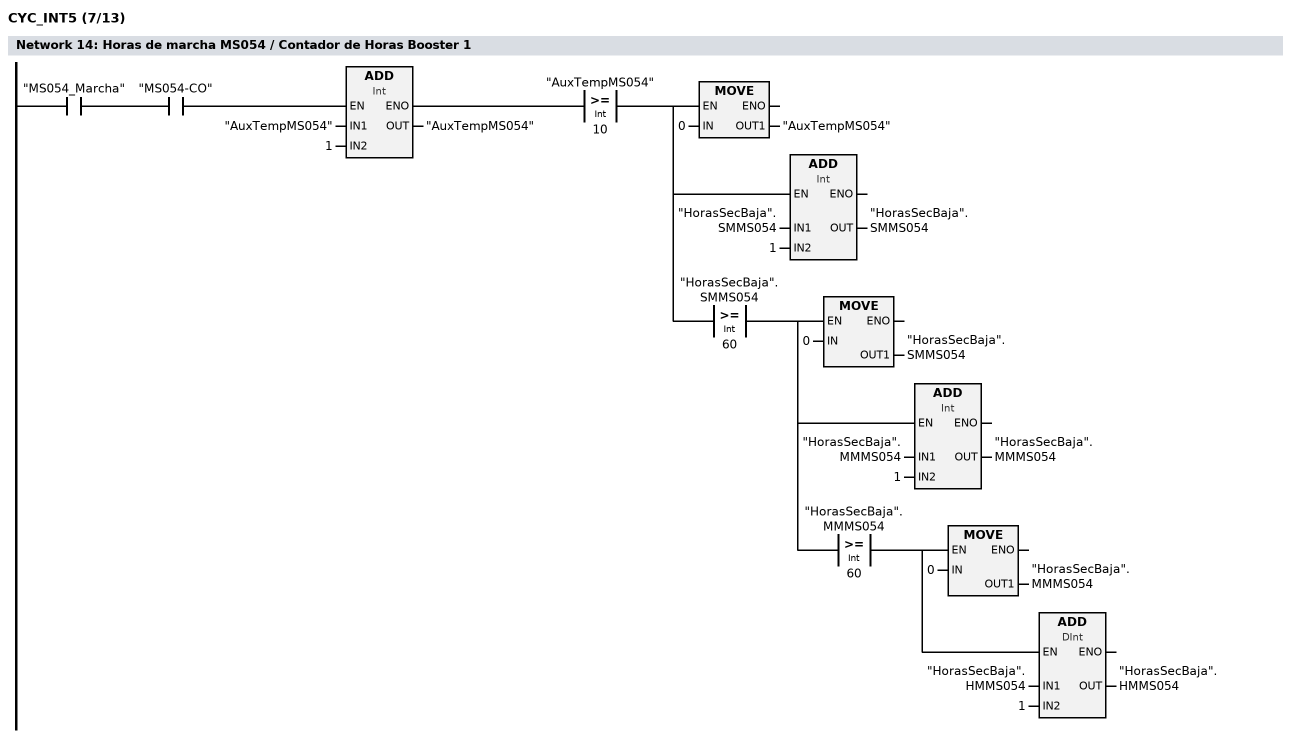
   RUNG wire#powerrail
      Contact( "MS054_Marcha" )
      Contact( "MS054-CO" )
      { S7_Templates := "SrcType := Int"; S7_GenerateENO := "TRUE" } Add(in1 := "AuxTempMS054", in2 := 1, out => "AuxTempMS054")
      { S7_Templates := "SrcType := Int" } GE_Contact(in1 := "AuxTempMS054", in2 := 10)
      wire#w1
      { S7_GenerateENO := "TRUE" } Move(in := 0, out1 => "AuxTempMS054")
   END_RUNG
   RUNG wire#w1
      { S7_Templates := "SrcType := Int"; S7_GenerateENO := "TRUE" } Add(in1 := "HorasSecBaja".SMMS054, in2 := 1, out => "HorasSecBaja".SMMS054)
   END_RUNG
   RUNG wire#w1
      { S7_Templates := "SrcType := Int" } GE_Contact(in1 := "HorasSecBaja".SMMS054, in2 := 60)
      wire#w2
      { S7_GenerateENO := "TRUE" } Move(in := 0, out1 => "HorasSecBaja".SMMS054)
   END_RUNG
   RUNG wire#w2
      { S7_Templates := "SrcType := Int"; S7_GenerateENO := "TRUE" } Add(in1 := "HorasSecBaja".MMMS054, in2 := 1, out => "HorasSecBaja".MMMS054)
   END_RUNG
   RUNG wire#w2
      { S7_Templates := "SrcType := Int" } GE_Contact(in1 := "HorasSecBaja".MMMS054, in2 := 60)
      wire#w3
      { S7_GenerateENO := "TRUE" } Move(in := 0, out1 => "HorasSecBaja".MMMS054)
   END_RUNG
   RUNG wire#w3
      { S7_Templates := "SrcType := DInt"; S7_GenerateENO := "TRUE" } Add(in1 := "HorasSecBaja".HMMS054, in2 := 1, out => "HorasSecBaja".HMMS054)
   END_RUNG
   // the same network as SCL:
   // ENO of a box is taken as its EN; it also drops when the box reports an error
   #_w1 := "MS054_Marcha" AND "MS054-CO";
   IF #_w1 THEN "AuxTempMS054" := "AuxTempMS054" + 1; END_IF;
   #_w2 := #_w1 AND ("AuxTempMS054" >= 10);
   IF #_w2 THEN
       "AuxTempMS054" := 0;
       "HorasSecBaja".SMMS054 := "HorasSecBaja".SMMS054 + 1;
   END_IF;
   #_w3 := #_w2 AND ("HorasSecBaja".SMMS054 >= 60);
   IF #_w3 THEN
       "HorasSecBaja".SMMS054 := 0;
       "HorasSecBaja".MMMS054 := "HorasSecBaja".MMMS054 + 1;
   END_IF;
   #_w4 := #_w3 AND ("HorasSecBaja".MMMS054 >= 60);
   IF #_w4 THEN
       "HorasSecBaja".MMMS054 := 0;
       "HorasSecBaja".HMMS054 := "HorasSecBaja".HMMS054 + 1;
   END_IF;
END_REGION

REGION Network 15: Horas de marcha MS055 / Contador de Horas Booster 1
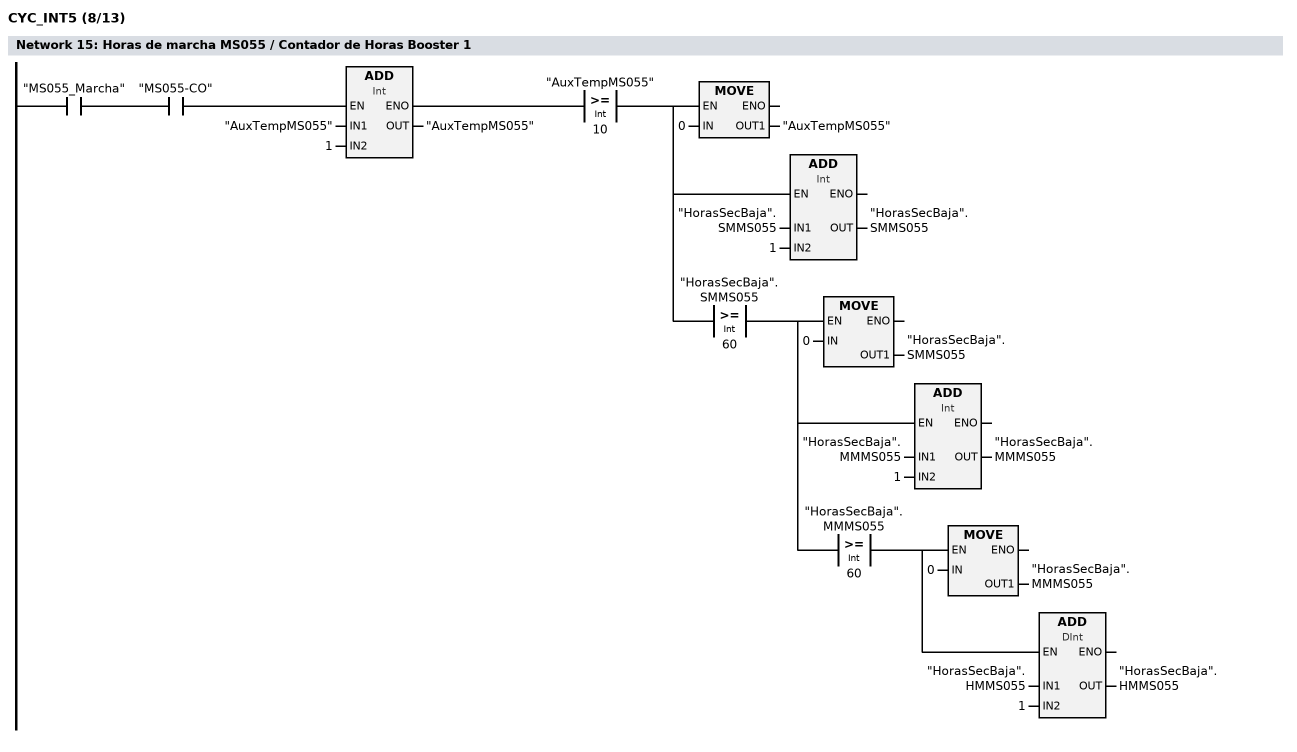
   RUNG wire#powerrail
      Contact( "MS055_Marcha" )
      Contact( "MS055-CO" )
      { S7_Templates := "SrcType := Int"; S7_GenerateENO := "TRUE" } Add(in1 := "AuxTempMS055", in2 := 1, out => "AuxTempMS055")
      { S7_Templates := "SrcType := Int" } GE_Contact(in1 := "AuxTempMS055", in2 := 10)
      wire#w1
      { S7_GenerateENO := "TRUE" } Move(in := 0, out1 => "AuxTempMS055")
   END_RUNG
   RUNG wire#w1
      { S7_Templates := "SrcType := Int"; S7_GenerateENO := "TRUE" } Add(in1 := "HorasSecBaja".SMMS055, in2 := 1, out => "HorasSecBaja".SMMS055)
   END_RUNG
   RUNG wire#w1
      { S7_Templates := "SrcType := Int" } GE_Contact(in1 := "HorasSecBaja".SMMS055, in2 := 60)
      wire#w2
      { S7_GenerateENO := "TRUE" } Move(in := 0, out1 => "HorasSecBaja".SMMS055)
   END_RUNG
   RUNG wire#w2
      { S7_Templates := "SrcType := Int"; S7_GenerateENO := "TRUE" } Add(in1 := "HorasSecBaja".MMMS055, in2 := 1, out => "HorasSecBaja".MMMS055)
   END_RUNG
   RUNG wire#w2
      { S7_Templates := "SrcType := Int" } GE_Contact(in1 := "HorasSecBaja".MMMS055, in2 := 60)
      wire#w3
      { S7_GenerateENO := "TRUE" } Move(in := 0, out1 => "HorasSecBaja".MMMS055)
   END_RUNG
   RUNG wire#w3
      { S7_Templates := "SrcType := DInt"; S7_GenerateENO := "TRUE" } Add(in1 := "HorasSecBaja".HMMS055, in2 := 1, out => "HorasSecBaja".HMMS055)
   END_RUNG
   // the same network as SCL:
   // ENO of a box is taken as its EN; it also drops when the box reports an error
   #_w1 := "MS055_Marcha" AND "MS055-CO";
   IF #_w1 THEN "AuxTempMS055" := "AuxTempMS055" + 1; END_IF;
   #_w2 := #_w1 AND ("AuxTempMS055" >= 10);
   IF #_w2 THEN
       "AuxTempMS055" := 0;
       "HorasSecBaja".SMMS055 := "HorasSecBaja".SMMS055 + 1;
   END_IF;
   #_w3 := #_w2 AND ("HorasSecBaja".SMMS055 >= 60);
   IF #_w3 THEN
       "HorasSecBaja".SMMS055 := 0;
       "HorasSecBaja".MMMS055 := "HorasSecBaja".MMMS055 + 1;
   END_IF;
   #_w4 := #_w3 AND ("HorasSecBaja".MMMS055 >= 60);
   IF #_w4 THEN
       "HorasSecBaja".MMMS055 := 0;
       "HorasSecBaja".HMMS055 := "HorasSecBaja".HMMS055 + 1;
   END_IF;
END_REGION

REGION Network 16: Horas de marcha MC060 / Contador de Horas Booster 1
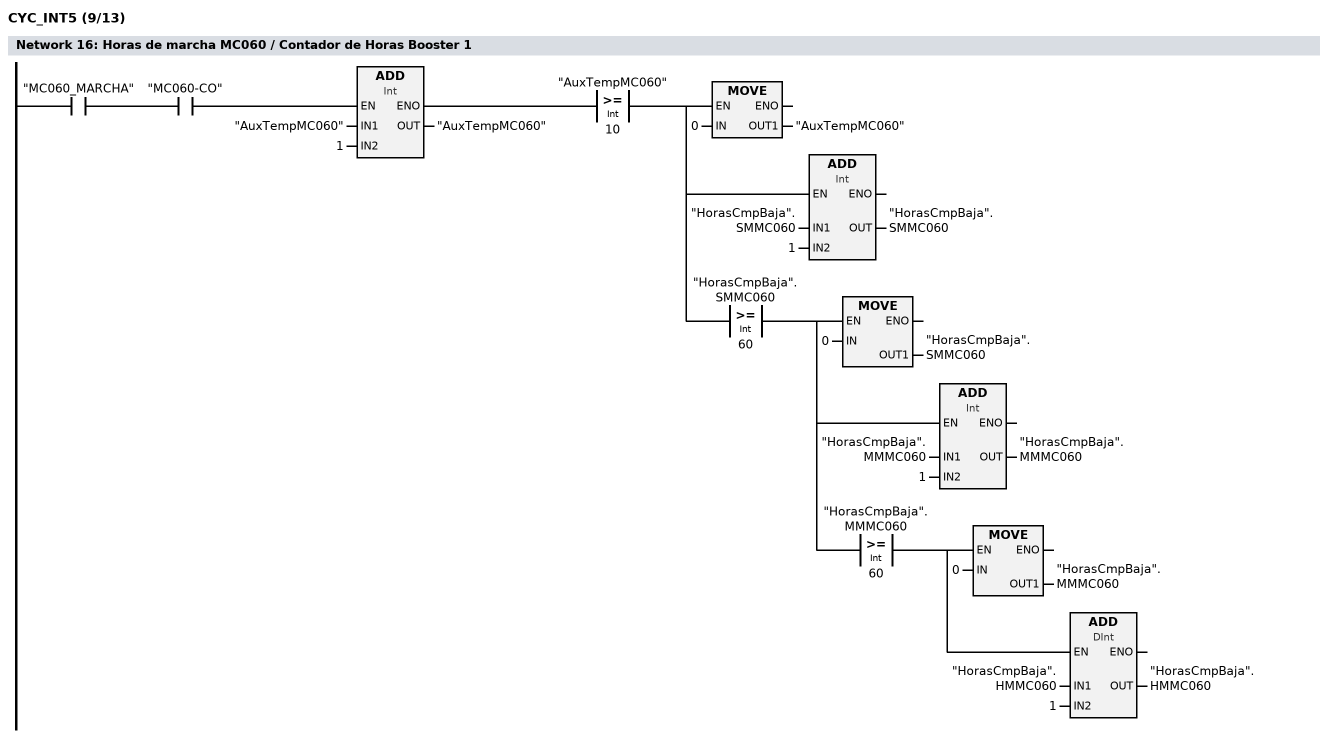
   RUNG wire#powerrail
      Contact( "MC060_MARCHA" )
      Contact( "MC060-CO" )
      { S7_Templates := "SrcType := Int"; S7_GenerateENO := "TRUE" } Add(in1 := "AuxTempMC060", in2 := 1, out => "AuxTempMC060")
      { S7_Templates := "SrcType := Int" } GE_Contact(in1 := "AuxTempMC060", in2 := 10)
      wire#w1
      { S7_GenerateENO := "TRUE" } Move(in := 0, out1 => "AuxTempMC060")
   END_RUNG
   RUNG wire#w1
      { S7_Templates := "SrcType := Int"; S7_GenerateENO := "TRUE" } Add(in1 := "HorasCmpBaja".SMMC060, in2 := 1, out => "HorasCmpBaja".SMMC060)
   END_RUNG
   RUNG wire#w1
      { S7_Templates := "SrcType := Int" } GE_Contact(in1 := "HorasCmpBaja".SMMC060, in2 := 60)
      wire#w2
      { S7_GenerateENO := "TRUE" } Move(in := 0, out1 => "HorasCmpBaja".SMMC060)
   END_RUNG
   RUNG wire#w2
      { S7_Templates := "SrcType := Int"; S7_GenerateENO := "TRUE" } Add(in1 := "HorasCmpBaja".MMMC060, in2 := 1, out => "HorasCmpBaja".MMMC060)
   END_RUNG
   RUNG wire#w2
      { S7_Templates := "SrcType := Int" } GE_Contact(in1 := "HorasCmpBaja".MMMC060, in2 := 60)
      wire#w3
      { S7_GenerateENO := "TRUE" } Move(in := 0, out1 => "HorasCmpBaja".MMMC060)
   END_RUNG
   RUNG wire#w3
      { S7_Templates := "SrcType := DInt"; S7_GenerateENO := "TRUE" } Add(in1 := "HorasCmpBaja".HMMC060, in2 := 1, out => "HorasCmpBaja".HMMC060)
   END_RUNG
   // the same network as SCL:
   // ENO of a box is taken as its EN; it also drops when the box reports an error
   #_w1 := "MC060_MARCHA" AND "MC060-CO";
   IF #_w1 THEN "AuxTempMC060" := "AuxTempMC060" + 1; END_IF;
   #_w2 := #_w1 AND ("AuxTempMC060" >= 10);
   IF #_w2 THEN
       "AuxTempMC060" := 0;
       "HorasCmpBaja".SMMC060 := "HorasCmpBaja".SMMC060 + 1;
   END_IF;
   #_w3 := #_w2 AND ("HorasCmpBaja".SMMC060 >= 60);
   IF #_w3 THEN
       "HorasCmpBaja".SMMC060 := 0;
       "HorasCmpBaja".MMMC060 := "HorasCmpBaja".MMMC060 + 1;
   END_IF;
   #_w4 := #_w3 AND ("HorasCmpBaja".MMMC060 >= 60);
   IF #_w4 THEN
       "HorasCmpBaja".MMMC060 := 0;
       "HorasCmpBaja".HMMC060 := "HorasCmpBaja".HMMC060 + 1;
   END_IF;
END_REGION

REGION Network 17: Horas de marcha MC061 / Contador de Horas Booster 1
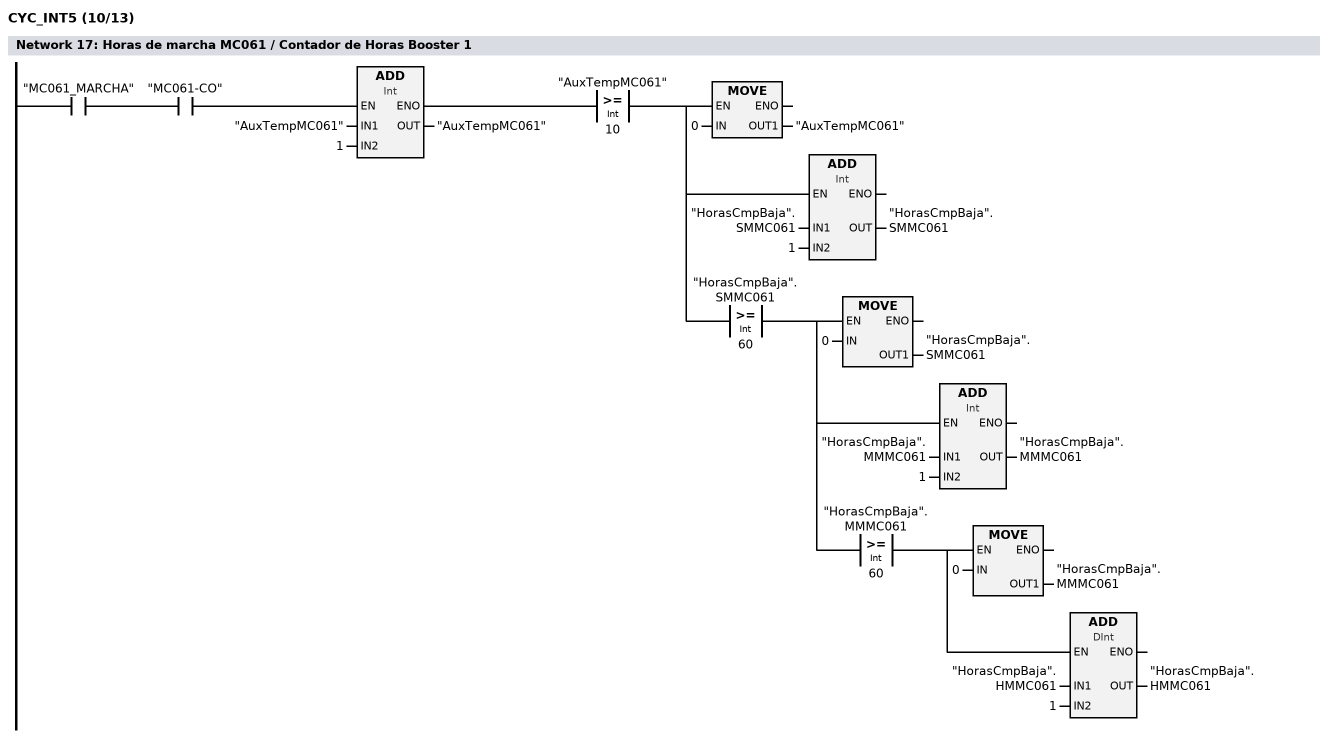
   RUNG wire#powerrail
      Contact( "MC061_MARCHA" )
      Contact( "MC061-CO" )
      { S7_Templates := "SrcType := Int"; S7_GenerateENO := "TRUE" } Add(in1 := "AuxTempMC061", in2 := 1, out => "AuxTempMC061")
      { S7_Templates := "SrcType := Int" } GE_Contact(in1 := "AuxTempMC061", in2 := 10)
      wire#w1
      { S7_GenerateENO := "TRUE" } Move(in := 0, out1 => "AuxTempMC061")
   END_RUNG
   RUNG wire#w1
      { S7_Templates := "SrcType := Int"; S7_GenerateENO := "TRUE" } Add(in1 := "HorasCmpBaja".SMMC061, in2 := 1, out => "HorasCmpBaja".SMMC061)
   END_RUNG
   RUNG wire#w1
      { S7_Templates := "SrcType := Int" } GE_Contact(in1 := "HorasCmpBaja".SMMC061, in2 := 60)
      wire#w2
      { S7_GenerateENO := "TRUE" } Move(in := 0, out1 => "HorasCmpBaja".SMMC061)
   END_RUNG
   RUNG wire#w2
      { S7_Templates := "SrcType := Int"; S7_GenerateENO := "TRUE" } Add(in1 := "HorasCmpBaja".MMMC061, in2 := 1, out => "HorasCmpBaja".MMMC061)
   END_RUNG
   RUNG wire#w2
      { S7_Templates := "SrcType := Int" } GE_Contact(in1 := "HorasCmpBaja".MMMC061, in2 := 60)
      wire#w3
      { S7_GenerateENO := "TRUE" } Move(in := 0, out1 => "HorasCmpBaja".MMMC061)
   END_RUNG
   RUNG wire#w3
      { S7_Templates := "SrcType := DInt"; S7_GenerateENO := "TRUE" } Add(in1 := "HorasCmpBaja".HMMC061, in2 := 1, out => "HorasCmpBaja".HMMC061)
   END_RUNG
   // the same network as SCL:
   // ENO of a box is taken as its EN; it also drops when the box reports an error
   #_w1 := "MC061_MARCHA" AND "MC061-CO";
   IF #_w1 THEN "AuxTempMC061" := "AuxTempMC061" + 1; END_IF;
   #_w2 := #_w1 AND ("AuxTempMC061" >= 10);
   IF #_w2 THEN
       "AuxTempMC061" := 0;
       "HorasCmpBaja".SMMC061 := "HorasCmpBaja".SMMC061 + 1;
   END_IF;
   #_w3 := #_w2 AND ("HorasCmpBaja".SMMC061 >= 60);
   IF #_w3 THEN
       "HorasCmpBaja".SMMC061 := 0;
       "HorasCmpBaja".MMMC061 := "HorasCmpBaja".MMMC061 + 1;
   END_IF;
   #_w4 := #_w3 AND ("HorasCmpBaja".MMMC061 >= 60);
   IF #_w4 THEN
       "HorasCmpBaja".MMMC061 := 0;
       "HorasCmpBaja".HMMC061 := "HorasCmpBaja".HMMC061 + 1;
   END_IF;
END_REGION

REGION Network 18: Horas de marcha MC062 / Contador de Horas Booster 1
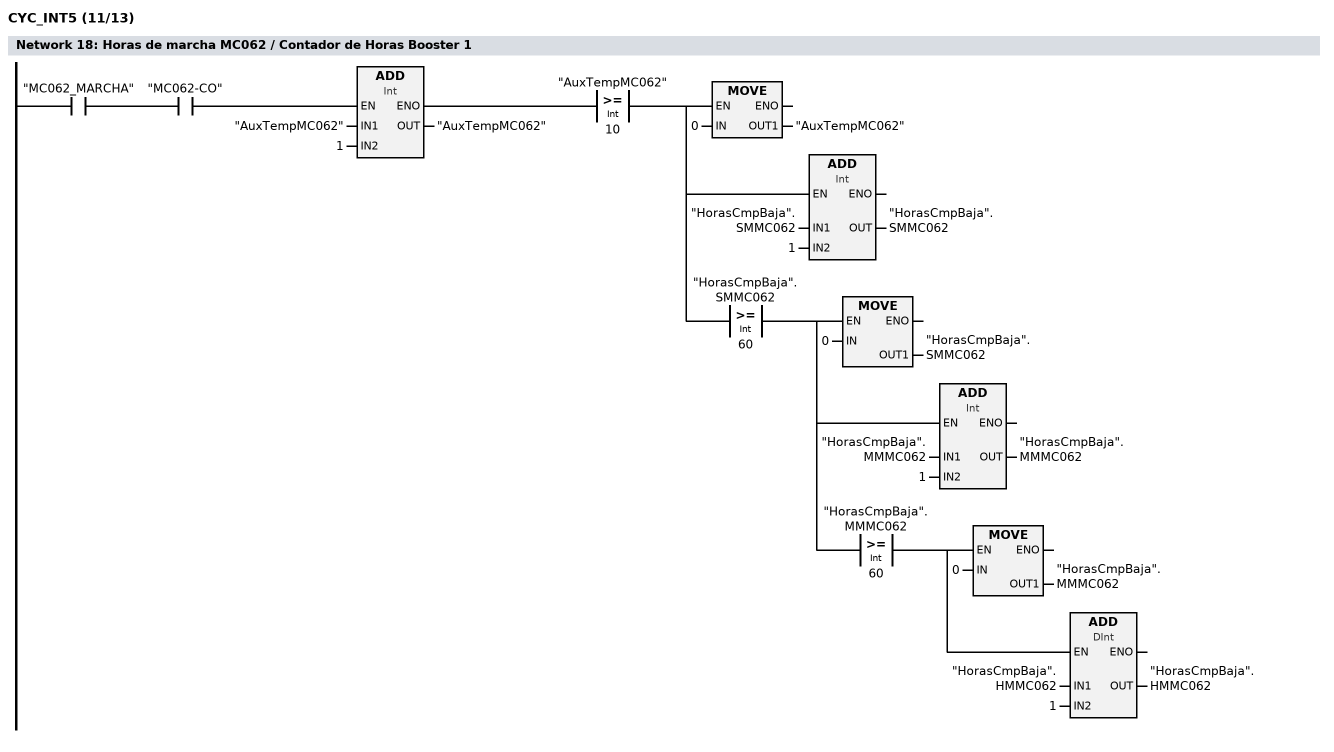
   RUNG wire#powerrail
      Contact( "MC062_MARCHA" )
      Contact( "MC062-CO" )
      { S7_Templates := "SrcType := Int"; S7_GenerateENO := "TRUE" } Add(in1 := "AuxTempMC062", in2 := 1, out => "AuxTempMC062")
      { S7_Templates := "SrcType := Int" } GE_Contact(in1 := "AuxTempMC062", in2 := 10)
      wire#w1
      { S7_GenerateENO := "TRUE" } Move(in := 0, out1 => "AuxTempMC062")
   END_RUNG
   RUNG wire#w1
      { S7_Templates := "SrcType := Int"; S7_GenerateENO := "TRUE" } Add(in1 := "HorasCmpBaja".SMMC062, in2 := 1, out => "HorasCmpBaja".SMMC062)
   END_RUNG
   RUNG wire#w1
      { S7_Templates := "SrcType := Int" } GE_Contact(in1 := "HorasCmpBaja".SMMC062, in2 := 60)
      wire#w2
      { S7_GenerateENO := "TRUE" } Move(in := 0, out1 => "HorasCmpBaja".SMMC062)
   END_RUNG
   RUNG wire#w2
      { S7_Templates := "SrcType := Int"; S7_GenerateENO := "TRUE" } Add(in1 := "HorasCmpBaja".MMMC062, in2 := 1, out => "HorasCmpBaja".MMMC062)
   END_RUNG
   RUNG wire#w2
      { S7_Templates := "SrcType := Int" } GE_Contact(in1 := "HorasCmpBaja".MMMC062, in2 := 60)
      wire#w3
      { S7_GenerateENO := "TRUE" } Move(in := 0, out1 => "HorasCmpBaja".MMMC062)
   END_RUNG
   RUNG wire#w3
      { S7_Templates := "SrcType := DInt"; S7_GenerateENO := "TRUE" } Add(in1 := "HorasCmpBaja".HMMC062, in2 := 1, out => "HorasCmpBaja".HMMC062)
   END_RUNG
   // the same network as SCL:
   // ENO of a box is taken as its EN; it also drops when the box reports an error
   #_w1 := "MC062_MARCHA" AND "MC062-CO";
   IF #_w1 THEN "AuxTempMC062" := "AuxTempMC062" + 1; END_IF;
   #_w2 := #_w1 AND ("AuxTempMC062" >= 10);
   IF #_w2 THEN
       "AuxTempMC062" := 0;
       "HorasCmpBaja".SMMC062 := "HorasCmpBaja".SMMC062 + 1;
   END_IF;
   #_w3 := #_w2 AND ("HorasCmpBaja".SMMC062 >= 60);
   IF #_w3 THEN
       "HorasCmpBaja".SMMC062 := 0;
       "HorasCmpBaja".MMMC062 := "HorasCmpBaja".MMMC062 + 1;
   END_IF;
   #_w4 := #_w3 AND ("HorasCmpBaja".MMMC062 >= 60);
   IF #_w4 THEN
       "HorasCmpBaja".MMMC062 := 0;
       "HorasCmpBaja".HMMC062 := "HorasCmpBaja".HMMC062 + 1;
   END_IF;
END_REGION

REGION Network 19: Horas de marcha MC063 / Contador de Horas Booster 1
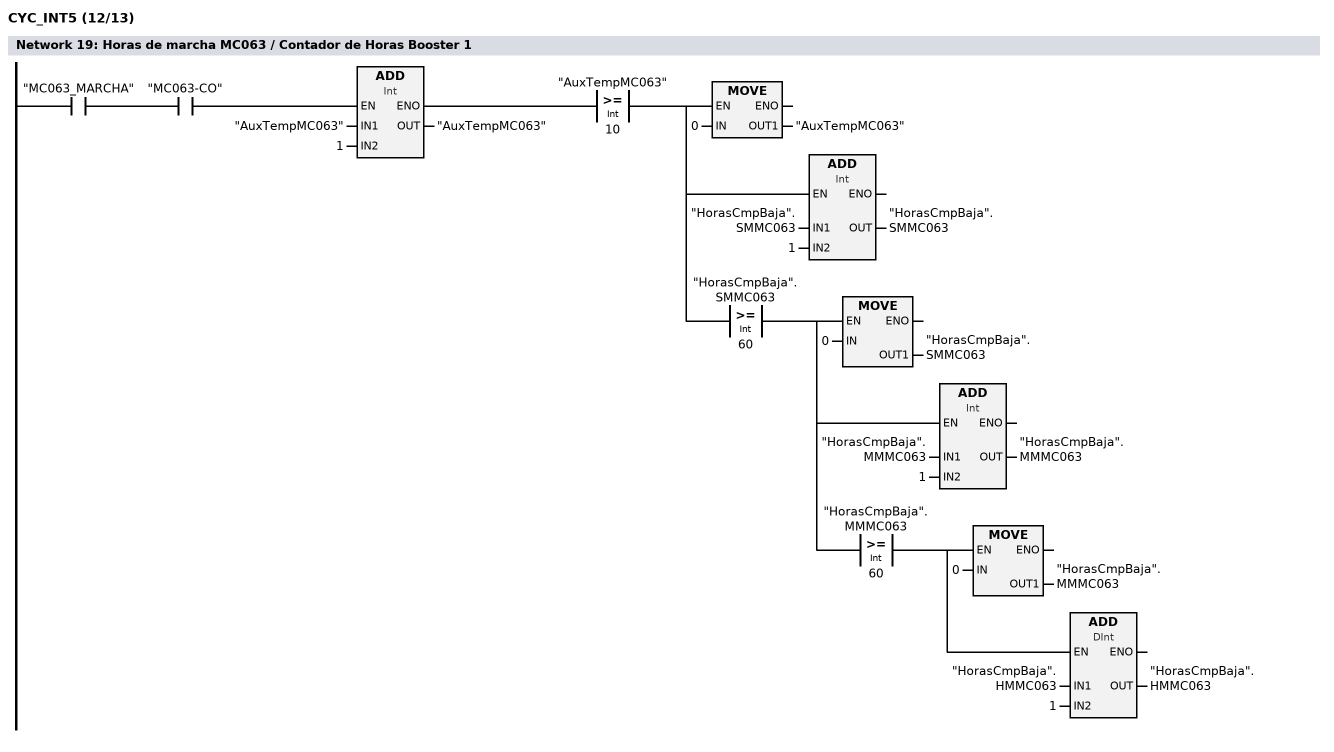
   RUNG wire#powerrail
      Contact( "MC063_MARCHA" )
      Contact( "MC063-CO" )
      { S7_Templates := "SrcType := Int"; S7_GenerateENO := "TRUE" } Add(in1 := "AuxTempMC063", in2 := 1, out => "AuxTempMC063")
      { S7_Templates := "SrcType := Int" } GE_Contact(in1 := "AuxTempMC063", in2 := 10)
      wire#w1
      { S7_GenerateENO := "TRUE" } Move(in := 0, out1 => "AuxTempMC063")
   END_RUNG
   RUNG wire#w1
      { S7_Templates := "SrcType := Int"; S7_GenerateENO := "TRUE" } Add(in1 := "HorasCmpBaja".SMMC063, in2 := 1, out => "HorasCmpBaja".SMMC063)
   END_RUNG
   RUNG wire#w1
      { S7_Templates := "SrcType := Int" } GE_Contact(in1 := "HorasCmpBaja".SMMC063, in2 := 60)
      wire#w2
      { S7_GenerateENO := "TRUE" } Move(in := 0, out1 => "HorasCmpBaja".SMMC063)
   END_RUNG
   RUNG wire#w2
      { S7_Templates := "SrcType := Int"; S7_GenerateENO := "TRUE" } Add(in1 := "HorasCmpBaja".MMMC063, in2 := 1, out => "HorasCmpBaja".MMMC063)
   END_RUNG
   RUNG wire#w2
      { S7_Templates := "SrcType := Int" } GE_Contact(in1 := "HorasCmpBaja".MMMC063, in2 := 60)
      wire#w3
      { S7_GenerateENO := "TRUE" } Move(in := 0, out1 => "HorasCmpBaja".MMMC063)
   END_RUNG
   RUNG wire#w3
      { S7_Templates := "SrcType := DInt"; S7_GenerateENO := "TRUE" } Add(in1 := "HorasCmpBaja".HMMC063, in2 := 1, out => "HorasCmpBaja".HMMC063)
   END_RUNG
   // the same network as SCL:
   // ENO of a box is taken as its EN; it also drops when the box reports an error
   #_w1 := "MC063_MARCHA" AND "MC063-CO";
   IF #_w1 THEN "AuxTempMC063" := "AuxTempMC063" + 1; END_IF;
   #_w2 := #_w1 AND ("AuxTempMC063" >= 10);
   IF #_w2 THEN
       "AuxTempMC063" := 0;
       "HorasCmpBaja".SMMC063 := "HorasCmpBaja".SMMC063 + 1;
   END_IF;
   #_w3 := #_w2 AND ("HorasCmpBaja".SMMC063 >= 60);
   IF #_w3 THEN
       "HorasCmpBaja".SMMC063 := 0;
       "HorasCmpBaja".MMMC063 := "HorasCmpBaja".MMMC063 + 1;
   END_IF;
   #_w4 := #_w3 AND ("HorasCmpBaja".MMMC063 >= 60);
   IF #_w4 THEN
       "HorasCmpBaja".MMMC063 := 0;
       "HorasCmpBaja".HMMC063 := "HorasCmpBaja".HMMC063 + 1;
   END_IF;
END_REGION

REGION Network 20: Horas de marcha MC064 / Contador de Horas Booster 1
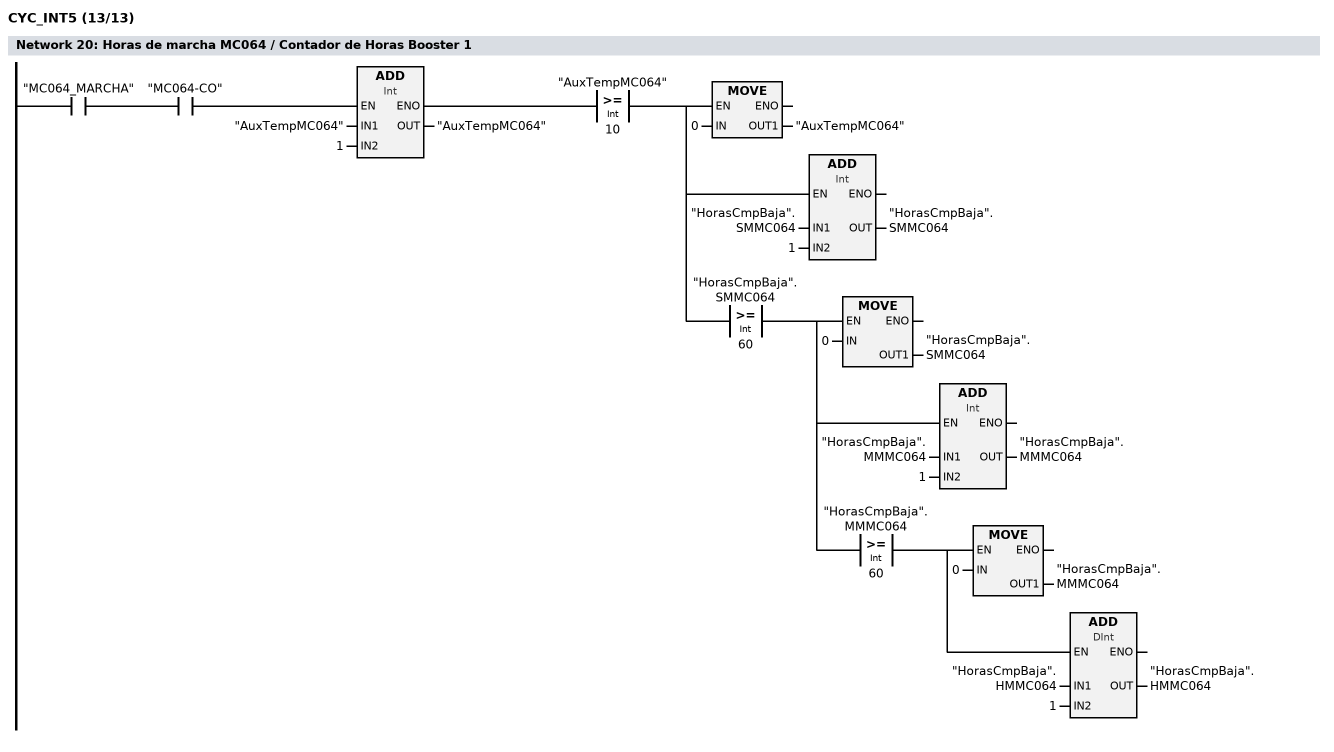
   RUNG wire#powerrail
      Contact( "MC064_MARCHA" )
      Contact( "MC064-CO" )
      { S7_Templates := "SrcType := Int"; S7_GenerateENO := "TRUE" } Add(in1 := "AuxTempMC064", in2 := 1, out => "AuxTempMC064")
      { S7_Templates := "SrcType := Int" } GE_Contact(in1 := "AuxTempMC064", in2 := 10)
      wire#w1
      { S7_GenerateENO := "TRUE" } Move(in := 0, out1 => "AuxTempMC064")
   END_RUNG
   RUNG wire#w1
      { S7_Templates := "SrcType := Int"; S7_GenerateENO := "TRUE" } Add(in1 := "HorasCmpBaja".SMMC064, in2 := 1, out => "HorasCmpBaja".SMMC064)
   END_RUNG
   RUNG wire#w1
      { S7_Templates := "SrcType := Int" } GE_Contact(in1 := "HorasCmpBaja".SMMC064, in2 := 60)
      wire#w2
      { S7_GenerateENO := "TRUE" } Move(in := 0, out1 => "HorasCmpBaja".SMMC064)
   END_RUNG
   RUNG wire#w2
      { S7_Templates := "SrcType := Int"; S7_GenerateENO := "TRUE" } Add(in1 := "HorasCmpBaja".MMMC064, in2 := 1, out => "HorasCmpBaja".MMMC064)
   END_RUNG
   RUNG wire#w2
      { S7_Templates := "SrcType := Int" } GE_Contact(in1 := "HorasCmpBaja".MMMC064, in2 := 60)
      wire#w3
      { S7_GenerateENO := "TRUE" } Move(in := 0, out1 => "HorasCmpBaja".MMMC064)
   END_RUNG
   RUNG wire#w3
      { S7_Templates := "SrcType := DInt"; S7_GenerateENO := "TRUE" } Add(in1 := "HorasCmpBaja".HMMC064, in2 := 1, out => "HorasCmpBaja".HMMC064)
   END_RUNG
   // the same network as SCL:
   // ENO of a box is taken as its EN; it also drops when the box reports an error
   #_w1 := "MC064_MARCHA" AND "MC064-CO";
   IF #_w1 THEN "AuxTempMC064" := "AuxTempMC064" + 1; END_IF;
   #_w2 := #_w1 AND ("AuxTempMC064" >= 10);
   IF #_w2 THEN
       "AuxTempMC064" := 0;
       "HorasCmpBaja".SMMC064 := "HorasCmpBaja".SMMC064 + 1;
   END_IF;
   #_w3 := #_w2 AND ("HorasCmpBaja".SMMC064 >= 60);
   IF #_w3 THEN
       "HorasCmpBaja".SMMC064 := 0;
       "HorasCmpBaja".MMMC064 := "HorasCmpBaja".MMMC064 + 1;
   END_IF;
   #_w4 := #_w3 AND ("HorasCmpBaja".MMMC064 >= 60);
   IF #_w4 THEN
       "HorasCmpBaja".MMMC064 := 0;
       "HorasCmpBaja".HMMC064 := "HorasCmpBaja".HMMC064 + 1;
   END_IF;
END_REGION
END_ORGANIZATION_BLOCK

// folder: OBs de Fallas

ORGANIZATION_BLOCK "OB40"   // OB40, STL
{ S7_Optimized_Access := 'FALSE' }
VERSION : 0.0
BEGIN
END_ORGANIZATION_BLOCK

ORGANIZATION_BLOCK "Cycle Time Fault"   // OB80, STL
{ S7_Optimized_Access := 'FALSE' }
VERSION : 0.0
BEGIN
END_ORGANIZATION_BLOCK

ORGANIZATION_BLOCK "I/O Point Fault 1"   // OB82, LAD
{ S7_Optimized_Access := 'FALSE' }
VERSION : 0.1
BEGIN
END_ORGANIZATION_BLOCK

ORGANIZATION_BLOCK "OB83"   // OB83, STL
{ S7_Optimized_Access := 'FALSE' }
VERSION : 0.1
BEGIN
END_ORGANIZATION_BLOCK

ORGANIZATION_BLOCK "OB Not Loaded Fault"   // OB85, LAD
{ S7_Optimized_Access := 'FALSE' }
VERSION : 0.1
BEGIN
END_ORGANIZATION_BLOCK

ORGANIZATION_BLOCK "Fallo del bastidor"   // OB86, STL
{ S7_Optimized_Access := 'FALSE' }
VERSION : 0.1
BEGIN
END_ORGANIZATION_BLOCK

ORGANIZATION_BLOCK "Communication Fault"   // OB87, LAD
{ S7_Optimized_Access := 'FALSE' }
VERSION : 0.1
BEGIN
END_ORGANIZATION_BLOCK

ORGANIZATION_BLOCK "Complete Restart"   // OB100, LAD
{ S7_Optimized_Access := 'FALSE' }
VERSION : 0.1
BEGIN
END_ORGANIZATION_BLOCK

ORGANIZATION_BLOCK "Programming Error"   // OB121, LAD
{ S7_Optimized_Access := 'FALSE' }
VERSION : 0.1
BEGIN
END_ORGANIZATION_BLOCK

ORGANIZATION_BLOCK "Module Access Error"   // OB122, LAD
{ S7_Optimized_Access := 'FALSE' }
VERSION : 0.1
BEGIN
END_ORGANIZATION_BLOCK

// folder: Panel

FUNCTION_BLOCK "CHControlMotorPanelMTA"   // FB55, LAD
{ S7_Optimized_Access := 'FALSE' }
VERSION : 0.1
   VAR_TEMP   // added for the SCL form of the ladder/FBD networks
      _w1 : Bool;
   END_VAR
BEGIN

REGION Network 1
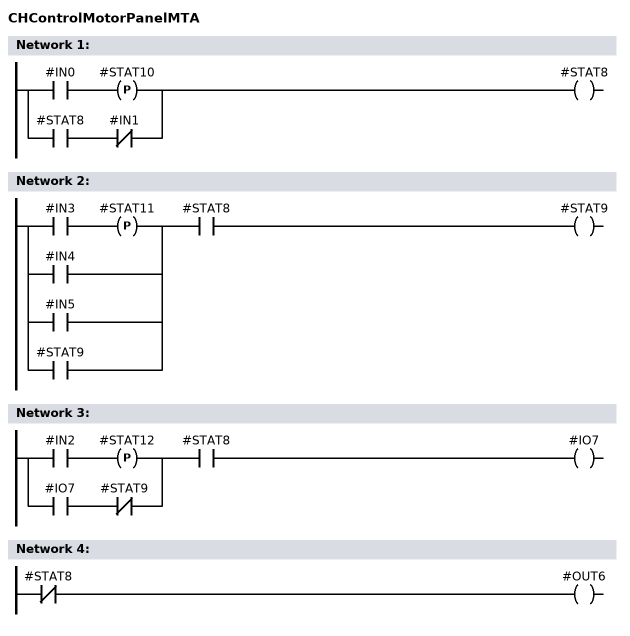
   RUNG wire#powerrail
      Contact( #IN0 )
      P_Trig( #STAT10 )
      wire#w1
      Coil( #STAT8 )
   END_RUNG
   RUNG wire#powerrail
      Contact( #STAT8 )
      I_Contact( #IN1 )
   END_RUNG wire#w1
   // the same network as SCL:
   #_w1 := #IN0 AND NOT #STAT10;   // rising edge
   #STAT10 := #IN0;
   #STAT8 := #_w1 OR (#STAT8 AND NOT #IN1);
END_REGION

REGION Network 2
   RUNG wire#powerrail
      Contact( #IN3 )
      P_Trig( #STAT11 )
      wire#w1
      Contact( #STAT8 )
      Coil( #STAT9 )
   END_RUNG
   RUNG wire#powerrail
      Contact( #IN4 )
   END_RUNG wire#w1
   RUNG wire#powerrail
      Contact( #IN5 )
   END_RUNG wire#w1
   RUNG wire#powerrail
      Contact( #STAT9 )
   END_RUNG wire#w1
   // the same network as SCL:
   #_w1 := #IN3 AND NOT #STAT11;   // rising edge
   #STAT11 := #IN3;
   #STAT9 := (#_w1 OR #IN4 OR #IN5 OR #STAT9) AND #STAT8;
END_REGION

REGION Network 3
   RUNG wire#powerrail
      Contact( #IN2 )
      P_Trig( #STAT12 )
      wire#w1
      Contact( #STAT8 )
      Coil( #IO7 )
   END_RUNG
   RUNG wire#powerrail
      Contact( #IO7 )
      I_Contact( #STAT9 )
   END_RUNG wire#w1
   // the same network as SCL:
   #_w1 := #IN2 AND NOT #STAT12;   // rising edge
   #STAT12 := #IN2;
   #IO7 := (#_w1 OR (#IO7 AND NOT #STAT9)) AND #STAT8;
END_REGION

REGION Network 4
   RUNG wire#powerrail
      I_Contact( #STAT8 )
      Coil( #OUT6 )
   END_RUNG
   // the same network as SCL:
   #OUT6 := NOT #STAT8;
END_REGION
END_FUNCTION_BLOCK

FUNCTION "AnimaciónMTA" : Void   // FC2, LAD
{ S7_Optimized_Access := 'FALSE' }
VERSION : 0.1
   VAR_TEMP   // added for the SCL form of the ladder/FBD networks
      _w1 : Bool;
      _w2 : Bool;
   END_VAR
BEGIN

REGION Network 1: Indicador Chillers
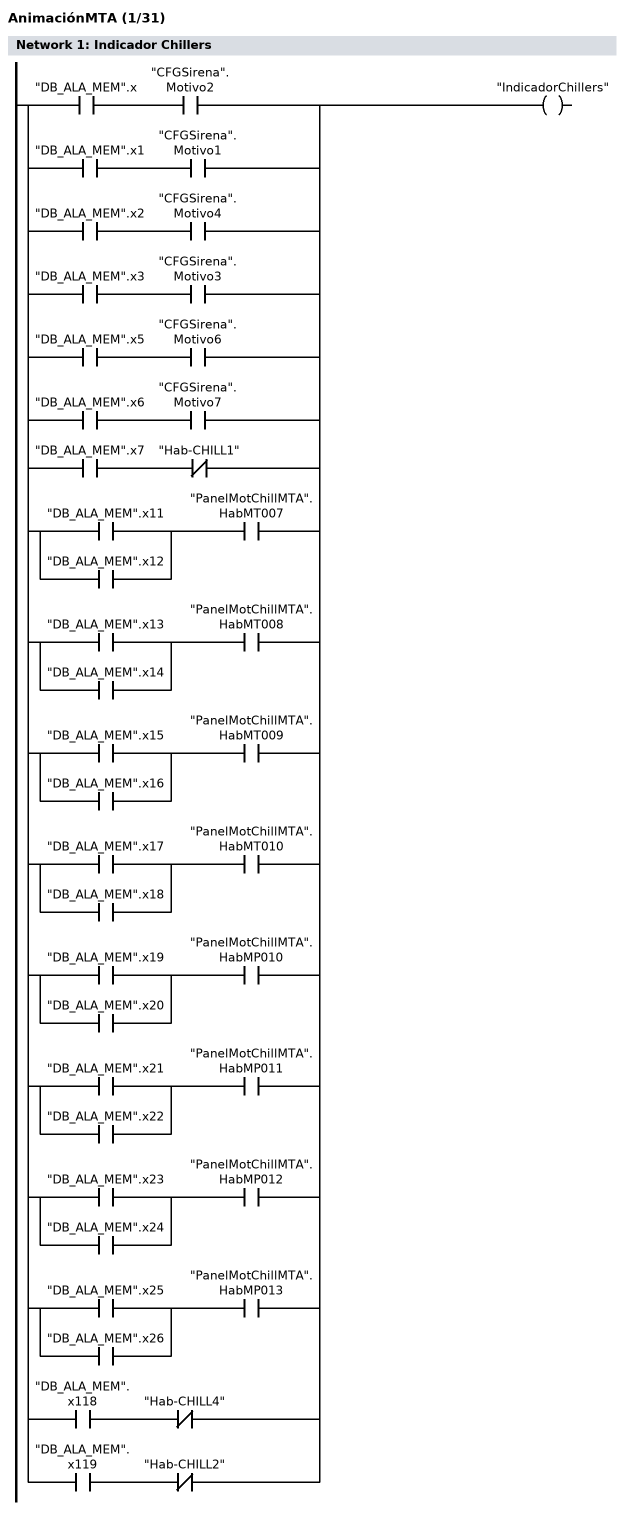
   RUNG wire#powerrail
      Contact( "DB_ALA_MEM".x )
      Contact( "CFGSirena".Motivo2 )
      wire#w1
      Coil( "IndicadorChillers" )
   END_RUNG
   RUNG wire#powerrail
      Contact( "DB_ALA_MEM".x1 )
      Contact( "CFGSirena".Motivo1 )
   END_RUNG wire#w1
   RUNG wire#powerrail
      Contact( "DB_ALA_MEM".x2 )
      Contact( "CFGSirena".Motivo4 )
   END_RUNG wire#w1
   RUNG wire#powerrail
      Contact( "DB_ALA_MEM".x3 )
      Contact( "CFGSirena".Motivo3 )
   END_RUNG wire#w1
   RUNG wire#powerrail
      Contact( "DB_ALA_MEM".x5 )
      Contact( "CFGSirena".Motivo6 )
   END_RUNG wire#w1
   RUNG wire#powerrail
      Contact( "DB_ALA_MEM".x6 )
      Contact( "CFGSirena".Motivo7 )
   END_RUNG wire#w1
   RUNG wire#powerrail
      Contact( "DB_ALA_MEM".x7 )
      I_Contact( "Hab-CHILL1" )
   END_RUNG wire#w1
   RUNG wire#powerrail
      Contact( "DB_ALA_MEM".x11 )
      wire#w2
      Contact( "PanelMotChillMTA".HabMT007 )
   END_RUNG wire#w1
   RUNG wire#powerrail
      Contact( "DB_ALA_MEM".x12 )
   END_RUNG wire#w2
   RUNG wire#powerrail
      Contact( "DB_ALA_MEM".x13 )
      wire#w3
      Contact( "PanelMotChillMTA".HabMT008 )
   END_RUNG wire#w1
   RUNG wire#powerrail
      Contact( "DB_ALA_MEM".x14 )
   END_RUNG wire#w3
   RUNG wire#powerrail
      Contact( "DB_ALA_MEM".x15 )
      wire#w4
      Contact( "PanelMotChillMTA".HabMT009 )
   END_RUNG wire#w1
   RUNG wire#powerrail
      Contact( "DB_ALA_MEM".x16 )
   END_RUNG wire#w4
   RUNG wire#powerrail
      Contact( "DB_ALA_MEM".x17 )
      wire#w5
      Contact( "PanelMotChillMTA".HabMT010 )
   END_RUNG wire#w1
   RUNG wire#powerrail
      Contact( "DB_ALA_MEM".x18 )
   END_RUNG wire#w5
   RUNG wire#powerrail
      Contact( "DB_ALA_MEM".x19 )
      wire#w6
      Contact( "PanelMotChillMTA".HabMP010 )
   END_RUNG wire#w1
   RUNG wire#powerrail
      Contact( "DB_ALA_MEM".x20 )
   END_RUNG wire#w6
   RUNG wire#powerrail
      Contact( "DB_ALA_MEM".x21 )
      wire#w7
      Contact( "PanelMotChillMTA".HabMP011 )
   END_RUNG wire#w1
   RUNG wire#powerrail
      Contact( "DB_ALA_MEM".x22 )
   END_RUNG wire#w7
   RUNG wire#powerrail
      Contact( "DB_ALA_MEM".x23 )
      wire#w8
      Contact( "PanelMotChillMTA".HabMP012 )
   END_RUNG wire#w1
   RUNG wire#powerrail
      Contact( "DB_ALA_MEM".x24 )
   END_RUNG wire#w8
   RUNG wire#powerrail
      Contact( "DB_ALA_MEM".x25 )
      wire#w9
      Contact( "PanelMotChillMTA".HabMP013 )
   END_RUNG wire#w1
   RUNG wire#powerrail
      Contact( "DB_ALA_MEM".x26 )
   END_RUNG wire#w9
   RUNG wire#powerrail
      Contact( "DB_ALA_MEM".x118 )
      I_Contact( "Hab-CHILL4" )
   END_RUNG wire#w1
   RUNG wire#powerrail
      Contact( "DB_ALA_MEM".x119 )
      I_Contact( "Hab-CHILL2" )
   END_RUNG wire#w1
   // the same network as SCL:
   "IndicadorChillers" := ("DB_ALA_MEM".x AND "CFGSirena".Motivo2) OR ("DB_ALA_MEM".x1 AND "CFGSirena".Motivo1) OR ("DB_ALA_MEM".x2 AND "CFGSirena".Motivo4) OR ("DB_ALA_MEM".x3 AND "CFGSirena".Motivo3) OR ("DB_ALA_MEM".x5 AND "CFGSirena".Motivo6) OR ("DB_ALA_MEM".x6 AND "CFGSirena".Motivo7) OR ("DB_ALA_MEM".x7 AND NOT "Hab-CHILL1") OR (("DB_ALA_MEM".x11 OR "DB_ALA_MEM".x12) AND "PanelMotChillMTA".HabMT007) OR (("DB_ALA_MEM".x13 OR "DB_ALA_MEM".x14) AND "PanelMotChillMTA".HabMT008) OR (("DB_ALA_MEM".x15 OR "DB_ALA_MEM".x16) AND "PanelMotChillMTA".HabMT009) OR (("DB_ALA_MEM".x17 OR "DB_ALA_MEM".x18) AND "PanelMotChillMTA".HabMT010) OR (("DB_ALA_MEM".x19 OR "DB_ALA_MEM".x20) AND "PanelMotChillMTA".HabMP010) OR (("DB_ALA_MEM".x21 OR "DB_ALA_MEM".x22) AND "PanelMotChillMTA".HabMP011) OR (("DB_ALA_MEM".x23 OR "DB_ALA_MEM".x24) AND "PanelMotChillMTA".HabMP012) OR (("DB_ALA_MEM".x25 OR "DB_ALA_MEM".x26) AND "PanelMotChillMTA".HabMP013) OR ("DB_ALA_MEM".x118 AND NOT "Hab-CHILL4") OR ("DB_ALA_MEM".x119 AND NOT "Hab-CHILL2");